
PopupScreen "Tank 1P Status" 885x425
   TrendView "Trend view_1" at 280,8 size 600x360
   TextField "Text field_4" at 20,136 size 86x22; Text 'Pressure:'
   IOField "I/O field_1" at 175,131 size 90x25; FormatPattern s999.9; Unit  mBar
      ProcessValue <- "20_TANKS_IP_DATA_RIO_01_FIRST_TANK_TANKS_PRESS"
   TextField "Text field_5" at 20,170 size 113x22; Text 'Water Level:'
   IOField "I/O field_2" at 175,165 size 90x25; FormatPattern 999.9; Unit  %
      ProcessValue <- "20_TANKS_IP_DATA_RIO_01_SECOND_TANK_BWT_LEVEL"
   TextField "Text field_6" at 20,204 size 137x22; Text 'MBG Flow Rate:'
   IOField "I/O field_3" at 175,199 size 90x25; FormatPattern 999.9; Unit  m³/hr
      ProcessValue <- "20_TANKS_IP_DATA_RIO_01_SECOND_TANK_MBG_FLOW"
   TextField "Text field_7" at 20,238 size 135x22; Text 'USD Flow Rate:'
   IOField "I/O field_4" at 175,233 size 90x25; FormatPattern 999.9; Unit  m³/hr
      ProcessValue <- "20_TANKS_IP_DATA_RIO_01_SECOND_TANK_USD_FLOW"
   TextField "Text field_8" at 20,272 size 140x22; Text 'Water pH Level:'
   IOField "I/O field_5" at 175,267 size 90x25; FormatPattern 99.9
      ProcessValue <- "20_TANKS_IP_DATA_RIO_01_SECOND_TANK_BWT_PH"
   TextField "Text field_9" at 20,306 size 143x22; Text 'Water DO Level:'
   IOField "I/O field_6" at 175,301 size 90x25; FormatPattern 99.99; Unit  mg/l
      ProcessValue <- "20_TANKS_IP_DATA_RIO_01_SECOND_TANK_BWT_DO"
   TextField "Text field_10" at 20,340 size 174x22; Text 'Water Temperature:'
   IOField "I/O field_7" at 190,335 size 75x25; FormatPattern 999.9; Unit  °C
      ProcessValue <- "20_TANKS_IP_DATA_RIO_01_SECOND_TANK_BWT_TEMP"
   Button "Button_1" at 51,5 size 219x35; TextOff 'Port Tank 1 (1P)'
      on Release: function_efd93a16("Tank 1P Status", 168, 315, -1, 0, 1)
   Button "Button_4" at 547,375 size 150x40; TextOff 'Disable Tank'; Authorization "Operate"
      on Press: function_b14e0dd5("504_Tank Grouping_DB2020_TANK ACTIV 2", 0)
   TextField "Text field_1" at 20,90 size 109x25; Text 'TIME LEFT:'
   GraphicView "Graphic view_1" at 20,46 size 245x32; Picture "Tank Manually Disabled"
   GraphicIOField "Graphic I/O field_1" at 20,46 size 245x32; PictureList "Tank Process Stage_II"
      ProcessValue <- "2110_BTCS_CNTRL_DB_BTCS_STATE"
      Visibility <- "504_Tank Grouping_DB2020_GROUP of TANK 2"
   Button "Button_2" at 4,5 size 45x35; TextOff 'Text'; PictureOff "Graphic_286"
      on Click: function_efd93a16("Tank 1P Status", 0, 0, -1, -1, 1)
   Button "Button_3" at 287,375 size 230x40; TextOff 'Text'; PictureList "Water Level Override"; Authorization "Operate"
      on Press: InvertBit("2062_Warning_Data_Water Level Override 1P")
      ProcessValue <- "2062_Warning_Data_Water Level Override 1P"
   Button "Button_5" at 27,375 size 230x40; TextOff 'Tank Shutdown Alarm'
      Visibility <- "2062_Warning_Data_Alarm Tank P1"
      ProcessValue <- "2062_Warning_Data_Water Level Override 1P"
   Button "Button_6" at 27,375 size 230x40; TextOff 'No/Low Water Level'; Authorization "Operate"
      Visibility <- "LT422 1P  TANK LEVEL ALARM_ALARM L"
      ProcessValue <- "2062_Warning_Data_Water Level Override 1P"
   IOField "I/O field_29" at 218,90 size 47x25; FormatPattern 99; Unit m
      ProcessValue <- "504_Tank Grouping_DB2020_Time Left Tank_Time Left m Tank 2"
   IOField "I/O field_8" at 173,90 size 42x25; FormatPattern 99; Unit h
      ProcessValue <- "504_Tank Grouping_DB2020_Time Left Tank_Time Left h Tank 2"
   IOField "I/O field_9" at 128,90 size 42x25; FormatPattern 99; Unit d
      ProcessValue <- "504_Tank Grouping_DB2020_Time Left Tank_Time Left d Tank 2"

PopupScreen "Tank 1S Status" 885x425
   TrendView "Trend view_1" at 280,7 size 600x360
   TextField "Text field_4" at 20,135 size 86x22; Text 'Pressure:'
   IOField "I/O field_1" at 175,130 size 90x25; FormatPattern s999.9; Unit  mBar
      ProcessValue <- "20_TANKS_IP_DATA_RIO_01_FIRST_TANK_TANKS_PRESS"
   TextField "Text field_5" at 20,169 size 113x22; Text 'Water Level:'
   IOField "I/O field_2" at 175,164 size 90x25; FormatPattern 999.9; Unit  %
      ProcessValue <- "20_TANKS_IP_DATA_RIO_01_THIRD_TANK_BWT_LEVEL"
   TextField "Text field_6" at 20,203 size 137x22; Text 'MBG Flow Rate:'
   IOField "I/O field_3" at 175,198 size 90x25; FormatPattern 999.9; Unit  m³/hr
      ProcessValue <- "20_TANKS_IP_DATA_RIO_01_THIRD_TANK_MBG_FLOW"
   TextField "Text field_7" at 20,237 size 135x22; Text 'USD Flow Rate:'
   IOField "I/O field_4" at 175,232 size 90x25; FormatPattern 999.9; Unit  m³/hr
      ProcessValue <- "20_TANKS_IP_DATA_RIO_01_THIRD_TANK_USD_FLOW"
   TextField "Text field_8" at 20,271 size 140x22; Text 'Water pH Level:'
   IOField "I/O field_5" at 175,266 size 90x25; FormatPattern 99.9
      ProcessValue <- "20_TANKS_IP_DATA_RIO_01_THIRD_TANK_BWT_PH"
   TextField "Text field_9" at 20,305 size 143x22; Text 'Water DO Level:'
   IOField "I/O field_6" at 175,300 size 90x25; FormatPattern 99.99; Unit  mg/l
      ProcessValue <- "20_TANKS_IP_DATA_RIO_01_THIRD_TANK_BWT_DO"
   TextField "Text field_10" at 20,339 size 174x22; Text 'Water Temperature:'
   IOField "I/O field_7" at 190,334 size 75x25; FormatPattern 999.9; Unit  °C
      ProcessValue <- "20_TANKS_IP_DATA_RIO_01_THIRD_TANK_BWT_TEMP"
   Button "Button_1" at 50,5 size 220x35; TextOff 'Starboard Tank 1 (1S)'
      on Release: function_efd93a16("Tank 1S Status", 168, 315, -1, 0, 1)
   Button "Button_4" at 548,375 size 150x40; TextOff 'Disable Tank'; Authorization "Operate"
      on Press: function_b14e0dd5("504_Tank Grouping_DB2020_TANK ACTIV 3", 0)
   TextField "Text field_1" at 20,90 size 109x25; Text 'TIME LEFT:'
   GraphicView "Graphic view_1" at 20,46 size 245x32; Picture "Tank Manually Disabled"
   GraphicIOField "Graphic I/O field_1" at 20,46 size 245x32; PictureList "Tank Process Stage_II"
      ProcessValue <- "2110_BTCS_CNTRL_DB_BTCS_STATE"
      Visibility <- "504_Tank Grouping_DB2020_GROUP of TANK 3"
   Button "Button_2" at 4,5 size 45x35; TextOff 'Text'; PictureOff "Graphic_286"
      on Click: function_efd93a16("Tank 1S Status", 0, 0, -1, -1, 1)
   Button "Button_3" at 287,375 size 230x40; TextOff 'Text'; PictureList "Water Level Override"; Authorization "Operate"
      on Press: InvertBit("2062_Warning_Data_Water Level Override 1S")
      ProcessValue <- "2062_Warning_Data_Water Level Override 1S"
   Button "Button_5" at 27,375 size 230x40; TextOff 'Tank Shutdown Alarm'
      Visibility <- "2062_Warning_Data_Alarm Tank S1"
   Button "Button_6" at 27,375 size 230x40; TextOff 'No/Low Water Level'; Authorization "Operate"
      Visibility <- "LT421 1S  TANK LEVEL ALARM_ALARM L"
   IOField "I/O field_29" at 218,90 size 47x25; FormatPattern 99; Unit m
      ProcessValue <- "504_Tank Grouping_DB2020_Time Left Tank_Time Left m Tank 3"
   IOField "I/O field_8" at 173,90 size 42x25; FormatPattern 99; Unit h
      ProcessValue <- "504_Tank Grouping_DB2020_Time Left Tank_Time Left h Tank 3"
   IOField "I/O field_9" at 128,90 size 42x25; FormatPattern 99; Unit d
      ProcessValue <- "504_Tank Grouping_DB2020_Time Left Tank_Time Left d Tank 3"

PopupScreen "Tank 2P Status" 885x425
   TrendView "Trend view_1" at 280,7 size 600x360
   TextField "Text field_4" at 20,135 size 86x22; Text 'Pressure:'
   IOField "I/O field_1" at 175,130 size 90x25; FormatPattern s999.9; Unit  mBar
      ProcessValue <- "20_TANKS_IP_DATA_RIO_02_FIRST_TANK_TANKS_PRESS"
   TextField "Text field_5" at 20,169 size 113x22; Text 'Water Level:'
   IOField "I/O field_2" at 175,164 size 90x25; FormatPattern 999.9; Unit  %
      ProcessValue <- "20_TANKS_IP_DATA_RIO_02_FIRST_TANK_BWT_LEVEL"
   TextField "Text field_6" at 20,203 size 137x22; Text 'MBG Flow Rate:'
   IOField "I/O field_3" at 175,198 size 90x25; FormatPattern 999.9; Unit  m³/hr
      ProcessValue <- "20_TANKS_IP_DATA_RIO_02_FIRST_TANK_MBG_FLOW"
   TextField "Text field_7" at 20,237 size 135x22; Text 'USD Flow Rate:'
   IOField "I/O field_4" at 175,232 size 90x25; FormatPattern 999.9; Unit  m³/hr
      ProcessValue <- "20_TANKS_IP_DATA_RIO_02_FIRST_TANK_USD_FLOW"
   TextField "Text field_8" at 20,271 size 140x22; Text 'Water pH Level:'
   IOField "I/O field_5" at 175,266 size 90x25; FormatPattern 99.9
      ProcessValue <- "20_TANKS_IP_DATA_RIO_02_FIRST_TANK_BWT_PH"
   TextField "Text field_9" at 20,305 size 143x22; Text 'Water DO Level:'
   IOField "I/O field_6" at 175,300 size 90x25; FormatPattern 99.99; Unit  mg/l
      ProcessValue <- "20_TANKS_IP_DATA_RIO_02_FIRST_TANK_BWT_DO"
   TextField "Text field_10" at 20,339 size 174x22; Text 'Water Temperature:'
   IOField "I/O field_7" at 190,334 size 75x25; FormatPattern 999.9; Unit  °C
      ProcessValue <- "20_TANKS_IP_DATA_RIO_02_FIRST_TANK_BWT_TEMP"
   Button "Button_4" at 545,375 size 150x40; TextOff 'Disable Tank'; Authorization "Operate"
      on Press: function_b14e0dd5("504_Tank Grouping_DB2020_TANK ACTIV 4", 0)
   Button "Button_1" at 51,5 size 219x35; TextOff 'Port Tank 2 (2P)'
      on Release: function_efd93a16("Tank 2P Status", 168, 315, -1, 0, 1)
   TextField "Text field_1" at 20,90 size 109x25; Text 'TIME LEFT:'
   GraphicView "Graphic view_1" at 20,46 size 245x32; Picture "Tank Manually Disabled"
   GraphicIOField "Graphic I/O field_1" at 20,46 size 245x32; PictureList "Tank Process Stage_II"
      ProcessValue <- "2110_BTCS_CNTRL_DB_BTCS_STATE"
      Visibility <- "504_Tank Grouping_DB2020_GROUP of TANK 4"
   Button "Button_2" at 4,5 size 45x35; TextOff 'Text'; PictureOff "Graphic_286"
      on Click: function_efd93a16("Tank 2P Status", 0, 0, -1, -1, 1)
   Button "Button_3" at 287,375 size 230x40; TextOff 'Text'; PictureList "Water Level Override"; Authorization "Operate"
      on Press: InvertBit("2062_Warning_Data_Water Level Override 2P")
      ProcessValue <- "2062_Warning_Data_Water Level Override 2P"
   Button "Button_5" at 27,375 size 230x40; TextOff 'Tank Shutdown Alarm'
      Visibility <- "2062_Warning_Data_Alarm Tank P2"
   Button "Button_6" at 27,375 size 230x40; TextOff 'No/Low Water Level'; Authorization "Operate"
      Visibility <- "FIT418_2P_ALM_ANALOG_DB_ALARM L"
   IOField "I/O field_29" at 218,90 size 47x25; FormatPattern 99; Unit m
      ProcessValue <- "504_Tank Grouping_DB2020_Time Left Tank_Time Left m Tank 4"
   IOField "I/O field_8" at 173,90 size 42x25; FormatPattern 99; Unit h
      ProcessValue <- "504_Tank Grouping_DB2020_Time Left Tank_Time Left h Tank 4"
   IOField "I/O field_9" at 128,90 size 42x25; FormatPattern 99; Unit d
      ProcessValue <- "504_Tank Grouping_DB2020_Time Left Tank_Time Left d Tank 4"

PopupScreen "Tank 2S Status" 885x425
   TrendView "Trend view_1" at 280,6 size 600x360
   TextField "Text field_4" at 20,134 size 86x22; Text 'Pressure:'
   IOField "I/O field_1" at 175,129 size 90x25; FormatPattern s999.9; Unit  mBar
      ProcessValue <- "20_TANKS_IP_DATA_RIO_02_FIRST_TANK_TANKS_PRESS"
   TextField "Text field_5" at 20,168 size 113x22; Text 'Water Level:'
   IOField "I/O field_2" at 175,163 size 90x25; FormatPattern 999.9; Unit  %
      ProcessValue <- "20_TANKS_IP_DATA_RIO_02_SECOND_TANK_BWT_LEVEL"
   TextField "Text field_6" at 20,202 size 137x22; Text 'MBG Flow Rate:'
   IOField "I/O field_3" at 175,197 size 90x25; FormatPattern 999.9; Unit  m³/hr
      ProcessValue <- "20_TANKS_IP_DATA_RIO_02_SECOND_TANK_MBG_FLOW"
   TextField "Text field_7" at 20,236 size 135x22; Text 'USD Flow Rate:'
   IOField "I/O field_4" at 175,231 size 90x25; FormatPattern 999.9; Unit  m³/hr
      ProcessValue <- "20_TANKS_IP_DATA_RIO_02_SECOND_TANK_USD_FLOW"
   TextField "Text field_8" at 20,270 size 140x22; Text 'Water pH Level:'
   IOField "I/O field_5" at 175,265 size 90x25; FormatPattern 99.9
      ProcessValue <- "20_TANKS_IP_DATA_RIO_02_SECOND_TANK_BWT_PH"
   TextField "Text field_9" at 20,304 size 143x22; Text 'Water DO Level:'
   IOField "I/O field_6" at 175,299 size 90x25; FormatPattern 99.99; Unit  mg/l
      ProcessValue <- "20_TANKS_IP_DATA_RIO_02_SECOND_TANK_BWT_DO"
   TextField "Text field_10" at 20,338 size 174x22; Text 'Water Temperature:'
   IOField "I/O field_7" at 190,333 size 75x25; FormatPattern 999.9; Unit  °C
      ProcessValue <- "20_TANKS_IP_DATA_RIO_02_SECOND_TANK_BWT_TEMP"
   Button "Button_4" at 550,375 size 150x40; TextOff 'Disable Tank'; Authorization "Operate"
      on Press: function_b14e0dd5("504_Tank Grouping_DB2020_TANK ACTIV 5", 0)
   Button "Button_1" at 50,5 size 220x35; TextOff 'Starboard Tank 2 (2S)'
      on Release: function_efd93a16("Tank 2S Status", 168, 315, -1, 0, 1)
   TextField "Text field_1" at 20,90 size 109x25; Text 'TIME LEFT:'
   GraphicView "Graphic view_1" at 20,46 size 245x32; Picture "Tank Manually Disabled"
   GraphicIOField "Graphic I/O field_1" at 20,46 size 245x32; PictureList "Tank Process Stage_II"
      ProcessValue <- "2110_BTCS_CNTRL_DB_BTCS_STATE"
      Visibility <- "504_Tank Grouping_DB2020_GROUP of TANK 5"
   Button "Button_2" at 4,5 size 45x35; TextOff 'Text'; PictureOff "Graphic_286"
      on Click: function_efd93a16("Tank 2S Status", 0, 0, -1, -1, 1)
   Button "Button_3" at 287,375 size 230x40; TextOff 'Text'; PictureList "Water Level Override"; Authorization "Operate"
      on Press: InvertBit("2062_Warning_Data_Water Level Override 2S")
      ProcessValue <- "2062_Warning_Data_Water Level Override 2S"
   Button "Button_5" at 27,375 size 230x40; TextOff 'Tank Shutdown Alarm'
      Visibility <- "2062_Warning_Data_Alarm Tank S2"
   Button "Button_6" at 27,375 size 230x40; TextOff 'No/Low Water Level'; Authorization "Operate"
      Visibility <- "LT421 2S  TANK LEVEL ALARM_ALARM L"
   IOField "I/O field_29" at 218,90 size 47x25; FormatPattern 99; Unit m
      ProcessValue <- "504_Tank Grouping_DB2020_Time Left Tank_Time Left m Tank 5"
   IOField "I/O field_8" at 173,90 size 42x25; FormatPattern 99; Unit h
      ProcessValue <- "504_Tank Grouping_DB2020_Time Left Tank_Time Left h Tank 5"
   IOField "I/O field_9" at 128,90 size 42x25; FormatPattern 99; Unit d
      ProcessValue <- "504_Tank Grouping_DB2020_Time Left Tank_Time Left d Tank 5"

PopupScreen "Tank 3P Status" 885x425
   TrendView "Trend view_1" at 280,7 size 600x360
   TextField "Text field_4" at 20,135 size 86x22; Text 'Pressure:'
   IOField "I/O field_1" at 175,130 size 90x25; FormatPattern s999.9; Unit  mBar
      ProcessValue <- "20_TANKS_IP_DATA_RIO_03_FIRST_TANK_TANKS_PRESS"
   TextField "Text field_5" at 20,169 size 113x22; Text 'Water Level:'
   IOField "I/O field_2" at 175,164 size 90x25; FormatPattern 999.9; Unit  %
      ProcessValue <- "20_TANKS_IP_DATA_RIO_03_FIRST_TANK_BWT_LEVEL"
   TextField "Text field_6" at 20,203 size 137x22; Text 'MBG Flow Rate:'
   IOField "I/O field_3" at 175,198 size 90x25; FormatPattern 999.9; Unit  m³/hr
      ProcessValue <- "20_TANKS_IP_DATA_RIO_03_FIRST_TANK_MBG_FLOW"
   TextField "Text field_7" at 20,237 size 135x22; Text 'USD Flow Rate:'
   IOField "I/O field_4" at 175,232 size 90x25; FormatPattern 999.9; Unit  m³/hr
      ProcessValue <- "20_TANKS_IP_DATA_RIO_03_FIRST_TANK_USD_FLOW"
   TextField "Text field_8" at 20,271 size 140x22; Text 'Water pH Level:'
   IOField "I/O field_5" at 175,266 size 90x25; FormatPattern 99.9
      ProcessValue <- "20_TANKS_IP_DATA_RIO_03_FIRST_TANK_BWT_PH"
   TextField "Text field_9" at 20,305 size 143x22; Text 'Water DO Level:'
   IOField "I/O field_6" at 175,300 size 90x25; FormatPattern 99.99; Unit  mg/l
      ProcessValue <- "20_TANKS_IP_DATA_RIO_03_FIRST_TANK_BWT_DO"
   TextField "Text field_10" at 20,339 size 174x22; Text 'Water Temperature:'
   IOField "I/O field_7" at 190,334 size 75x25; FormatPattern 999.9; Unit  °C
      ProcessValue <- "20_TANKS_IP_DATA_RIO_03_FIRST_TANK_BWT_TEMP"
   Button "Button_4" at 545,375 size 150x40; TextOff 'Disable Tank'; Authorization "Operate"
      on Press: function_b14e0dd5("504_Tank Grouping_DB2020_TANK ACTIV 6", 0)
   Button "Button_1" at 51,5 size 220x35; TextOff 'Port Tank 3 (3P)'
      on Release: function_efd93a16("Tank 3P Status", 168, 315, -1, 0, 1)
   TextField "Text field_1" at 20,90 size 109x25; Text 'TIME LEFT:'
   GraphicView "Graphic view_1" at 20,46 size 245x32; Picture "Tank Manually Disabled"
   GraphicIOField "Graphic I/O field_1" at 20,46 size 245x32; PictureList "Tank Process Stage_II"
      ProcessValue <- "2110_BTCS_CNTRL_DB_BTCS_STATE"
      Visibility <- "504_Tank Grouping_DB2020_GROUP of TANK 6"
   Button "Button_2" at 4,5 size 45x35; TextOff 'Text'; PictureOff "Graphic_286"
      on Click: function_efd93a16("Tank 3P Status", 0, 0, -1, -1, 1)
   Button "Button_3" at 287,375 size 230x40; TextOff 'Text'; PictureList "Water Level Override"; Authorization "Operate"
      on Press: InvertBit("2062_Warning_Data_Water Level Override 3P")
      ProcessValue <- "2062_Warning_Data_Water Level Override 3P"
   Button "Button_5" at 27,375 size 230x40; TextOff 'Tank Shutdown Alarm'
      Visibility <- "2062_Warning_Data_Alarm Tank P3"
   Button "Button_6" at 27,375 size 230x40; TextOff 'No/Low Water Level'; Authorization "Operate"
      Visibility <- "LT422 3P  TANK LEVEL ALARM_ALARM L"
   IOField "I/O field_29" at 218,90 size 47x25; FormatPattern 99; Unit m
      ProcessValue <- "504_Tank Grouping_DB2020_Time Left Tank_Time Left m Tank 6"
   IOField "I/O field_8" at 173,90 size 42x25; FormatPattern 99; Unit h
      ProcessValue <- "504_Tank Grouping_DB2020_Time Left Tank_Time Left h Tank 6"
   IOField "I/O field_9" at 128,90 size 42x25; FormatPattern 99; Unit d
      ProcessValue <- "504_Tank Grouping_DB2020_Time Left Tank_Time Left d Tank 6"

PopupScreen "Tank 3S Status" 885x425
   TrendView "Trend view_1" at 280,7 size 600x360
   TextField "Text field_4" at 20,135 size 86x22; Text 'Pressure:'
   IOField "I/O field_1" at 175,130 size 90x25; FormatPattern s999.9; Unit  mBar
      ProcessValue <- "20_TANKS_IP_DATA_RIO_03_FIRST_TANK_TANKS_PRESS"
   TextField "Text field_5" at 20,169 size 113x22; Text 'Water Level:'
   IOField "I/O field_2" at 175,164 size 90x25; FormatPattern 999.9; Unit  %
      ProcessValue <- "20_TANKS_IP_DATA_RIO_03_SECOND_TANK_BWT_LEVEL"
   TextField "Text field_6" at 20,203 size 137x22; Text 'MBG Flow Rate:'
   IOField "I/O field_3" at 175,198 size 90x25; FormatPattern 999.9; Unit  m³/hr
      ProcessValue <- "20_TANKS_IP_DATA_RIO_03_SECOND_TANK_MBG_FLOW"
   TextField "Text field_7" at 20,237 size 135x22; Text 'USD Flow Rate:'
   IOField "I/O field_4" at 175,232 size 90x25; FormatPattern 999.9; Unit  m³/hr
      ProcessValue <- "20_TANKS_IP_DATA_RIO_03_SECOND_TANK_USD_FLOW"
   TextField "Text field_8" at 20,271 size 140x22; Text 'Water pH Level:'
   IOField "I/O field_5" at 175,266 size 90x25; FormatPattern 99.9
      ProcessValue <- "20_TANKS_IP_DATA_RIO_03_SECOND_TANK_BWT_PH"
   TextField "Text field_9" at 20,305 size 143x22; Text 'Water DO Level:'
   IOField "I/O field_6" at 175,300 size 90x25; FormatPattern 99.99; Unit  mg/l
      ProcessValue <- "20_TANKS_IP_DATA_RIO_03_SECOND_TANK_BWT_DO"
   TextField "Text field_10" at 20,339 size 174x22; Text 'Water Temperature:'
   IOField "I/O field_7" at 190,334 size 75x25; FormatPattern 999.9; Unit  °C
      ProcessValue <- "20_TANKS_IP_DATA_RIO_03_SECOND_TANK_BWT_TEMP"
   Button "Button_4" at 547,375 size 150x40; TextOff 'Disable Tank'; Authorization "Operate"
      on Press: function_b14e0dd5("504_Tank Grouping_DB2020_TANK ACTIV 7", 0)
   Button "Button_1" at 51,5 size 219x35; TextOff 'Starboard Tank 3 (3S)'
      on Release: function_efd93a16("Tank 3S Status", 168, 315, -1, 0, 1)
   TextField "Text field_1" at 20,90 size 109x25; Text 'TIME LEFT:'
   GraphicView "Graphic view_1" at 20,46 size 245x32; Picture "Tank Manually Disabled"
   GraphicIOField "Graphic I/O field_1" at 20,46 size 245x32; PictureList "Tank Process Stage_II"
      ProcessValue <- "2110_BTCS_CNTRL_DB_BTCS_STATE"
      Visibility <- "504_Tank Grouping_DB2020_GROUP of TANK 7"
   Button "Button_2" at 4,5 size 45x35; TextOff 'Text'; PictureOff "Graphic_286"
      on Click: function_efd93a16("Tank 3S Status", 0, 0, -1, -1, 1)
   Button "Button_3" at 287,375 size 230x40; TextOff 'Text'; PictureList "Water Level Override"; Authorization "Operate"
      on Press: InvertBit("2062_Warning_Data_Water Level Override 3S")
      ProcessValue <- "2062_Warning_Data_Water Level Override 3S"
   Button "Button_5" at 27,375 size 230x40; TextOff 'Tank Shutdown Alarm'
      Visibility <- "2062_Warning_Data_Alarm Tank S3"
   Button "Button_6" at 27,375 size 230x40; TextOff 'No/Low Water Level'; Authorization "Operate"
      Visibility <- "LT421 3S  TANK LEVEL ALARM_ALARM L"
   IOField "I/O field_29" at 218,90 size 47x25; FormatPattern 99; Unit m
      ProcessValue <- "504_Tank Grouping_DB2020_Time Left Tank_Time Left m Tank 7"
   IOField "I/O field_8" at 173,90 size 42x25; FormatPattern 99; Unit h
      ProcessValue <- "504_Tank Grouping_DB2020_Time Left Tank_Time Left h Tank 7"
   IOField "I/O field_9" at 128,90 size 42x25; FormatPattern 99; Unit d
      ProcessValue <- "504_Tank Grouping_DB2020_Time Left Tank_Time Left d Tank 7"

PopupScreen "Tank 4P Status" 885x425
   TrendView "Trend view_1" at 280,7 size 600x360
   TextField "Text field_4" at 20,135 size 86x22; Text 'Pressure:'
   IOField "I/O field_1" at 175,130 size 90x25; FormatPattern s999.9; Unit  mBar
      ProcessValue <- "20_TANKS_IP_DATA_RIO_04_FIRST_TANK_TANKS_PRESS"
   TextField "Text field_5" at 20,169 size 113x22; Text 'Water Level:'
   IOField "I/O field_2" at 175,164 size 90x25; FormatPattern 999.9; Unit  %
      ProcessValue <- "20_TANKS_IP_DATA_RIO_04_FIRST_TANK_BWT_LEVEL"
   TextField "Text field_6" at 20,203 size 137x22; Text 'MBG Flow Rate:'
   IOField "I/O field_3" at 175,198 size 90x25; FormatPattern 999.9; Unit  m³/hr
      ProcessValue <- "20_TANKS_IP_DATA_RIO_04_FIRST_TANK_MBG_FLOW"
   TextField "Text field_7" at 20,237 size 135x22; Text 'USD Flow Rate:'
   IOField "I/O field_4" at 175,232 size 90x25; FormatPattern 999.9; Unit  m³/hr
      ProcessValue <- "20_TANKS_IP_DATA_RIO_04_FIRST_TANK_USD_FLOW"
   TextField "Text field_8" at 20,271 size 140x22; Text 'Water pH Level:'
   IOField "I/O field_5" at 175,266 size 90x25; FormatPattern 99.9
      ProcessValue <- "20_TANKS_IP_DATA_RIO_04_FIRST_TANK_BWT_PH"
   TextField "Text field_9" at 20,305 size 143x22; Text 'Water DO Level:'
   IOField "I/O field_6" at 175,300 size 90x25; FormatPattern 99.99; Unit  mg/l
      ProcessValue <- "20_TANKS_IP_DATA_RIO_04_FIRST_TANK_BWT_DO"
   TextField "Text field_10" at 20,339 size 174x22; Text 'Water Temperature:'
   IOField "I/O field_7" at 190,334 size 75x25; FormatPattern 999.9; Unit  °C
      ProcessValue <- "20_TANKS_IP_DATA_RIO_04_FIRST_TANK_BWT_TEMP"
   Button "Button_4" at 545,375 size 150x40; TextOff 'Disable Tank'; Authorization "Operate"
      on Press: function_b14e0dd5("504_Tank Grouping_DB2020_TANK ACTIV 8", 0)
   Button "Button_1" at 51,5 size 219x35; TextOff 'Port Tank 4 (4P)'
      on Release: function_efd93a16("Tank 4P Status", 168, 315, -1, 2, 1)
   TextField "Text field_1" at 20,90 size 109x25; Text 'TIME LEFT:'
   GraphicView "Graphic view_1" at 20,46 size 245x32; Picture "Tank Manually Disabled"
   GraphicIOField "Graphic I/O field_1" at 20,46 size 245x32; PictureList "Tank Process Stage_II"
      ProcessValue <- "2110_BTCS_CNTRL_DB_BTCS_STATE"
      Visibility <- "504_Tank Grouping_DB2020_GROUP of TANK 8"
   Button "Button_2" at 4,5 size 45x35; TextOff 'Text'; PictureOff "Graphic_286"
      on Click: function_efd93a16("Tank 4P Status", 0, 0, -1, -1, 1)
   Button "Button_3" at 287,375 size 230x40; TextOff 'Text'; PictureList "Water Level Override"; Authorization "Operate"
      on Press: InvertBit("2062_Warning_Data_Water Level Override 4P")
      ProcessValue <- "2062_Warning_Data_Water Level Override 4P"
   Button "Button_5" at 27,375 size 230x40; TextOff 'Tank Shutdown Alarm'
      Visibility <- "2062_Warning_Data_Alarm Tank P4"
   Button "Button_6" at 27,375 size 230x40; TextOff 'No/Low Water Level'; Authorization "Operate"
      Visibility <- "LT422 4P  TANK LEVEL ALARM_ALARM L"
   IOField "I/O field_29" at 218,90 size 47x25; FormatPattern 99; Unit m
      ProcessValue <- "504_Tank Grouping_DB2020_Time Left Tank_Time Left m Tank 8"
   IOField "I/O field_8" at 173,90 size 42x25; FormatPattern 99; Unit h
      ProcessValue <- "504_Tank Grouping_DB2020_Time Left Tank_Time Left h Tank 8"
   IOField "I/O field_9" at 128,90 size 42x25; FormatPattern 99; Unit d
      ProcessValue <- "504_Tank Grouping_DB2020_Time Left Tank_Time Left d Tank 8"

PopupScreen "Tank 4S Status" 885x425
   TrendView "Trend view_1" at 280,7 size 600x360
   TextField "Text field_4" at 20,135 size 86x22; Text 'Pressure:'
   IOField "I/O field_1" at 175,130 size 90x25; FormatPattern s999.9; Unit  mBar
      ProcessValue <- "20_TANKS_IP_DATA_RIO_04_FIRST_TANK_TANKS_PRESS"
   TextField "Text field_5" at 20,169 size 113x22; Text 'Water Level:'
   IOField "I/O field_2" at 175,164 size 90x25; FormatPattern 999.9; Unit  %
      ProcessValue <- "20_TANKS_IP_DATA_RIO_04_SECOND_TANK_BWT_LEVEL"
   TextField "Text field_6" at 20,203 size 137x22; Text 'MBG Flow Rate:'
   IOField "I/O field_3" at 175,198 size 90x25; FormatPattern 999.9; Unit  m³/hr
      ProcessValue <- "20_TANKS_IP_DATA_RIO_04_SECOND_TANK_MBG_FLOW"
   TextField "Text field_7" at 20,237 size 135x22; Text 'USD Flow Rate:'
   IOField "I/O field_4" at 175,232 size 90x25; FormatPattern 999.9; Unit  m³/hr
      ProcessValue <- "20_TANKS_IP_DATA_RIO_04_SECOND_TANK_USD_FLOW"
   TextField "Text field_8" at 20,271 size 140x22; Text 'Water pH Level:'
   IOField "I/O field_5" at 175,266 size 90x25; FormatPattern 99.9
      ProcessValue <- "20_TANKS_IP_DATA_RIO_04_SECOND_TANK_BWT_PH"
   TextField "Text field_9" at 20,305 size 143x22; Text 'Water DO Level:'
   IOField "I/O field_6" at 175,300 size 90x25; FormatPattern 99.99; Unit  mg/l
      ProcessValue <- "20_TANKS_IP_DATA_RIO_04_SECOND_TANK_BWT_DO"
   TextField "Text field_10" at 20,339 size 174x22; Text 'Water Temperature:'
   IOField "I/O field_7" at 190,334 size 75x25; FormatPattern 999.9; Unit  °C
      ProcessValue <- "20_TANKS_IP_DATA_RIO_04_SECOND_TANK_BWT_TEMP"
   Button "Button_4" at 545,375 size 150x40; TextOff 'Disable Tank'; Authorization "Operate"
      on Press: function_b14e0dd5("504_Tank Grouping_DB2020_TANK ACTIV 9", 0)
   Button "Button_1" at 50,5 size 220x35; TextOff 'Starboard Tank 4 (4S)'
      on Release: function_efd93a16("Tank 4S Status", 168, 315, -1, 2, 1)
   TextField "Text field_1" at 20,90 size 109x25; Text 'TIME LEFT:'
   GraphicView "Graphic view_1" at 20,46 size 245x32; Picture "Tank Manually Disabled"
   GraphicIOField "Graphic I/O field_1" at 20,46 size 245x32; PictureList "Tank Process Stage_II"
      ProcessValue <- "2110_BTCS_CNTRL_DB_BTCS_STATE"
      Visibility <- "504_Tank Grouping_DB2020_GROUP of TANK 9"
   Button "Button_2" at 4,5 size 45x35; TextOff 'Text'; PictureOff "Graphic_286"
      on Click: function_efd93a16("Tank 4S Status", 0, 0, -1, -1, 1)
   Button "Button_3" at 287,375 size 230x40; TextOff 'Text'; PictureList "Water Level Override"; Authorization "Operate"
      on Press: InvertBit("2062_Warning_Data_Water Level Override 4S")
      ProcessValue <- "2062_Warning_Data_Water Level Override 4S"
   Button "Button_5" at 27,375 size 230x40; TextOff 'Tank Shutdown Alarm'
      Visibility <- "2062_Warning_Data_Alarm Tank S4"
   Button "Button_6" at 27,375 size 230x40; TextOff 'No/Low Water Level'; Authorization "Operate"
      Visibility <- "LT421 4S  TANK LEVEL ALARM_ALARM L"
   IOField "I/O field_29" at 218,90 size 47x25; FormatPattern 99; Unit m
      ProcessValue <- "504_Tank Grouping_DB2020_Time Left Tank_Time Left m Tank 9"
   IOField "I/O field_8" at 173,90 size 42x25; FormatPattern 99; Unit h
      ProcessValue <- "504_Tank Grouping_DB2020_Time Left Tank_Time Left h Tank 9"
   IOField "I/O field_9" at 128,90 size 42x25; FormatPattern 99; Unit d
      ProcessValue <- "504_Tank Grouping_DB2020_Time Left Tank_Time Left d Tank 9"

PopupScreen "Tank 5P Status" 885x425
   TrendView "Trend view_1" at 280,7 size 600x360
   TextField "Text field_4" at 20,135 size 86x22; Text 'Pressure:'
   IOField "I/O field_1" at 175,130 size 90x25; FormatPattern s999.9; Unit  mBar
      ProcessValue <- "20_TANKS_IP_DATA_RIO_05_FIRST_TANK_TANKS_PRESS"
   TextField "Text field_5" at 20,169 size 113x22; Text 'Water Level:'
   IOField "I/O field_2" at 175,164 size 90x25; FormatPattern 999.9; Unit  %
      ProcessValue <- "20_TANKS_IP_DATA_RIO_05_FIRST_TANK_BWT_LEVEL"
   TextField "Text field_6" at 20,203 size 137x22; Text 'MBG Flow Rate:'
   IOField "I/O field_3" at 175,198 size 90x25; FormatPattern 999.9; Unit  m³/hr
      ProcessValue <- "20_TANKS_IP_DATA_RIO_05_FIRST_TANK_MBG_FLOW"
   TextField "Text field_7" at 20,237 size 135x22; Text 'USD Flow Rate:'
   IOField "I/O field_4" at 175,232 size 90x25; FormatPattern 999.9; Unit  m³/hr
      ProcessValue <- "20_TANKS_IP_DATA_RIO_05_FIRST_TANK_USD_FLOW"
   TextField "Text field_8" at 20,271 size 140x22; Text 'Water pH Level:'
   IOField "I/O field_5" at 175,266 size 90x25; FormatPattern 99.9
      ProcessValue <- "20_TANKS_IP_DATA_RIO_05_FIRST_TANK_BWT_PH"
   TextField "Text field_9" at 20,305 size 143x22; Text 'Water DO Level:'
   IOField "I/O field_6" at 175,300 size 90x25; FormatPattern 99.99; Unit  mg/l
      ProcessValue <- "20_TANKS_IP_DATA_RIO_05_FIRST_TANK_BWT_DO"
   TextField "Text field_10" at 20,339 size 174x22; Text 'Water Temperature:'
   IOField "I/O field_7" at 190,334 size 75x25; FormatPattern 999.9; Unit  °C
      ProcessValue <- "20_TANKS_IP_DATA_RIO_05_FIRST_TANK_BWT_TEMP"
   Button "Button_4" at 546,375 size 150x40; TextOff 'Disable Tank'; Authorization "Operate"
      on Press: function_b14e0dd5("504_Tank Grouping_DB2020_TANK ACTIV 10", 0)
   Button "Button_1" at 51,5 size 219x35; TextOff 'Port Tank 5 (5P)'
      on Release: function_efd93a16("Tank 5P Status", 168, 315, -1, 2, 1)
   TextField "Text field_1" at 20,90 size 109x25; Text 'TIME LEFT:'
   GraphicView "Graphic view_1" at 20,46 size 245x32; Picture "Tank Manually Disabled"
   GraphicIOField "Graphic I/O field_1" at 20,46 size 245x32; PictureList "Tank Process Stage_II"
      ProcessValue <- "2110_BTCS_CNTRL_DB_BTCS_STATE"
      Visibility <- "504_Tank Grouping_DB2020_GROUP of TANK 10"
   Button "Button_2" at 4,5 size 45x35; TextOff 'Text'; PictureOff "Graphic_286"
      on Click: function_efd93a16("Tank 5P Status", 0, 0, -1, -1, 1)
   Button "Button_3" at 287,375 size 230x40; TextOff 'Text'; PictureList "Water Level Override"; Authorization "Operate"
      on Press: InvertBit("2062_Warning_Data_Water Level Override 5P")
      ProcessValue <- "2062_Warning_Data_Water Level Override 5P"
   Button "Button_5" at 27,375 size 230x40; TextOff 'Tank Shutdown Alarm'
      Visibility <- "2062_Warning_Data_Alarm Tank P5"
   Button "Button_6" at 27,375 size 230x40; TextOff 'No/Low Water Level'; Authorization "Operate"
      Visibility <- "LT422 5P  TANK LEVEL ALARM_ALARM L"
   IOField "I/O field_29" at 218,90 size 47x25; FormatPattern 99; Unit m
      ProcessValue <- "504_Tank Grouping_DB2020_Time Left Tank_Time Left m Tank 10"
   IOField "I/O field_8" at 173,90 size 42x25; FormatPattern 99; Unit h
      ProcessValue <- "504_Tank Grouping_DB2020_Time Left Tank_Time Left h Tank 10"
   IOField "I/O field_9" at 128,90 size 42x25; FormatPattern 99; Unit d
      ProcessValue <- "504_Tank Grouping_DB2020_Time Left Tank_Time Left d Tank 10"

PopupScreen "Tank 5S Status" 885x425
   TrendView "Trend view_1" at 280,7 size 600x360
   TextField "Text field_4" at 20,135 size 86x22; Text 'Pressure:'
   IOField "I/O field_1" at 175,130 size 90x25; FormatPattern s999.9; Unit  mBar
      ProcessValue <- "20_TANKS_IP_DATA_RIO_05_FIRST_TANK_TANKS_PRESS"
   TextField "Text field_5" at 20,169 size 113x22; Text 'Water Level:'
   IOField "I/O field_2" at 175,164 size 90x25; FormatPattern 999.9; Unit  %
      ProcessValue <- "20_TANKS_IP_DATA_RIO_05_SECOND_TANK_BWT_LEVEL"
   TextField "Text field_6" at 20,203 size 137x22; Text 'MBG Flow Rate:'
   IOField "I/O field_3" at 175,198 size 90x25; FormatPattern 999.9; Unit  m³/hr
      ProcessValue <- "20_TANKS_IP_DATA_RIO_05_SECOND_TANK_MBG_FLOW"
   TextField "Text field_7" at 20,237 size 135x22; Text 'USD Flow Rate:'
   IOField "I/O field_4" at 175,232 size 90x25; FormatPattern 999.9; Unit  m³/hr
      ProcessValue <- "20_TANKS_IP_DATA_RIO_05_SECOND_TANK_USD_FLOW"
   TextField "Text field_8" at 20,271 size 140x22; Text 'Water pH Level:'
   IOField "I/O field_5" at 175,266 size 90x25; FormatPattern 99.9
      ProcessValue <- "20_TANKS_IP_DATA_RIO_05_SECOND_TANK_BWT_PH"
   TextField "Text field_9" at 20,305 size 143x22; Text 'Water DO Level:'
   IOField "I/O field_6" at 175,300 size 90x25; FormatPattern 99.99; Unit  mg/l
      ProcessValue <- "20_TANKS_IP_DATA_RIO_05_SECOND_TANK_BWT_DO"
   TextField "Text field_10" at 20,339 size 174x22; Text 'Water Temperature:'
   IOField "I/O field_7" at 190,334 size 75x25; FormatPattern 999.9; Unit  °C
      ProcessValue <- "20_TANKS_IP_DATA_RIO_05_SECOND_TANK_BWT_TEMP"
   Button "Button_4" at 550,375 size 150x40; TextOff 'Disable Tank'; Authorization "Operate"
      on Press: function_b14e0dd5("504_Tank Grouping_DB2020_TANK ACTIV 11", 0)
   Button "Button_1" at 50,5 size 220x35; TextOff 'Starboard Tank 5 (5S)'
      on Release: function_efd93a16("Tank 5S Status", 168, 315, -1, 2, 1)
   TextField "Text field_1" at 20,90 size 109x25; Text 'TIME LEFT:'
   GraphicView "Graphic view_1" at 20,46 size 245x32; Picture "Tank Manually Disabled"
   GraphicIOField "Graphic I/O field_1" at 20,46 size 245x32; PictureList "Tank Process Stage_II"
      ProcessValue <- "2110_BTCS_CNTRL_DB_BTCS_STATE"
      Visibility <- "504_Tank Grouping_DB2020_GROUP of TANK 11"
   Button "Button_2" at 4,5 size 45x35; TextOff 'Text'; PictureOff "Graphic_286"
      on Click: function_efd93a16("Tank 5S Status", 0, 0, -1, -1, 1)
   Button "Button_3" at 287,375 size 230x40; TextOff 'Text'; PictureList "Water Level Override"; Authorization "Operate"
      on Press: InvertBit("2062_Warning_Data_Water Level Override 5S")
      ProcessValue <- "2062_Warning_Data_Water Level Override 5S"
   Button "Button_5" at 27,375 size 230x40; TextOff 'Tank Shutdown Alarm'
      Visibility <- "2062_Warning_Data_Alarm Tank S5"
   Button "Button_6" at 27,375 size 230x40; TextOff 'No/Low Water Level'; Authorization "Operate"
      Visibility <- "LT421 5S  TANK LEVEL ALARM_ALARM L"
   IOField "I/O field_29" at 218,90 size 47x25; FormatPattern 99; Unit m
      ProcessValue <- "504_Tank Grouping_DB2020_Time Left Tank_Time Left m Tank 11"
   IOField "I/O field_8" at 173,90 size 42x25; FormatPattern 99; Unit h
      ProcessValue <- "504_Tank Grouping_DB2020_Time Left Tank_Time Left h Tank 11"
   IOField "I/O field_9" at 128,90 size 42x25; FormatPattern 99; Unit d
      ProcessValue <- "504_Tank Grouping_DB2020_Time Left Tank_Time Left d Tank 11"

PopupScreen "Tank 6P Status" 885x425
   TrendView "Trend view_1" at 280,7 size 600x360
   TextField "Text field_4" at 20,135 size 86x22; Text 'Pressure:'
   IOField "I/O field_1" at 175,130 size 90x25; FormatPattern s999.9; Unit  mBar
      ProcessValue <- "20_TANKS_IP_DATA_RIO_06_FIRST_TANK_TANKS_PRESS"
   TextField "Text field_5" at 20,169 size 113x22; Text 'Water Level:'
   IOField "I/O field_2" at 175,164 size 90x25; FormatPattern 999.9; Unit  %
      ProcessValue <- "20_TANKS_IP_DATA_RIO_06_FIRST_TANK_BWT_LEVEL"
   TextField "Text field_6" at 20,203 size 137x22; Text 'MBG Flow Rate:'
   IOField "I/O field_3" at 175,198 size 90x25; FormatPattern 999.9; Unit  m³/hr
      ProcessValue <- "20_TANKS_IP_DATA_RIO_06_FIRST_TANK_MBG_FLOW"
   TextField "Text field_7" at 20,237 size 135x22; Text 'USD Flow Rate:'
   IOField "I/O field_4" at 175,232 size 90x25; FormatPattern 999.9; Unit  m³/hr
      ProcessValue <- "20_TANKS_IP_DATA_RIO_06_FIRST_TANK_USD_FLOW"
   TextField "Text field_8" at 20,271 size 140x22; Text 'Water pH Level:'
   IOField "I/O field_5" at 175,266 size 90x25; FormatPattern 99.9
      ProcessValue <- "20_TANKS_IP_DATA_RIO_06_FIRST_TANK_BWT_PH"
   TextField "Text field_9" at 20,305 size 143x22; Text 'Water DO Level:'
   IOField "I/O field_6" at 175,300 size 90x25; FormatPattern 99.99; Unit  mg/l
      ProcessValue <- "20_TANKS_IP_DATA_RIO_06_FIRST_TANK_BWT_DO"
   TextField "Text field_10" at 20,339 size 174x22; Text 'Water Temperature:'
   IOField "I/O field_7" at 190,334 size 75x25; FormatPattern 999.9; Unit  °C
      ProcessValue <- "20_TANKS_IP_DATA_RIO_06_FIRST_TANK_BWT_TEMP"
   Button "Button_4" at 542,374 size 150x40; TextOff 'Disable Tank'; Authorization "Operate"
      on Press: function_b14e0dd5("504_Tank Grouping_DB2020_TANK ACTIV 12", 0)
   Button "Button_1" at 51,5 size 219x35; TextOff 'Port Tank 6 (6P)'
      on Release: function_efd93a16("Tank 6P Status", 168, 315, -1, 2, 1)
   TextField "Text field_1" at 20,90 size 109x25; Text 'TIME LEFT:'
   GraphicView "Graphic view_1" at 20,46 size 245x32; Picture "Tank Manually Disabled"
   GraphicIOField "Graphic I/O field_1" at 20,46 size 245x32; PictureList "Tank Process Stage_II"
      ProcessValue <- "2110_BTCS_CNTRL_DB_BTCS_STATE"
      Visibility <- "504_Tank Grouping_DB2020_GROUP of TANK 12"
   Button "Button_2" at 4,5 size 45x35; TextOff 'Text'; PictureOff "Graphic_286"
      on Click: function_efd93a16("Tank 6P Status", 0, 0, -1, -1, 1)
   Button "Button_3" at 287,375 size 230x40; TextOff 'Text'; PictureList "Water Level Override"; Authorization "Operate"
      on Press: InvertBit("2062_Warning_Data_Water Level Override 6P")
      ProcessValue <- "2062_Warning_Data_Water Level Override 6P"
   Button "Button_5" at 27,375 size 230x40; TextOff 'Tank Shutdown Alarm'
      Visibility <- "2062_Warning_Data_Alarm Tank P6"
   Button "Button_6" at 27,375 size 230x40; TextOff 'No/Low Water Level'; Authorization "Operate"
      Visibility <- "LT422 6P  TANK LEVEL ALARM_ALARM L"
   IOField "I/O field_29" at 218,90 size 47x25; FormatPattern 99; Unit m
      ProcessValue <- "504_Tank Grouping_DB2020_Time Left Tank_Time Left m Tank 12"
   IOField "I/O field_8" at 173,90 size 42x25; FormatPattern 99; Unit h
      ProcessValue <- "504_Tank Grouping_DB2020_Time Left Tank_Time Left h Tank 12"
   IOField "I/O field_9" at 128,90 size 42x25; FormatPattern 99; Unit d
      ProcessValue <- "504_Tank Grouping_DB2020_Time Left Tank_Time Left d Tank 12"

PopupScreen "Tank 6S Status" 885x425
   TrendView "Trend view_1" at 280,7 size 600x360
   TextField "Text field_4" at 20,135 size 86x22; Text 'Pressure:'
   IOField "I/O field_1" at 175,130 size 90x25; FormatPattern s999.9; Unit  mBar
      ProcessValue <- "20_TANKS_IP_DATA_RIO_06_FIRST_TANK_TANKS_PRESS"
   TextField "Text field_5" at 20,169 size 113x22; Text 'Water Level:'
   IOField "I/O field_2" at 175,164 size 90x25; FormatPattern 999.9; Unit  %
      ProcessValue <- "20_TANKS_IP_DATA_RIO_06_SECOND_TANK_BWT_LEVEL"
   TextField "Text field_6" at 20,203 size 137x22; Text 'MBG Flow Rate:'
   IOField "I/O field_3" at 175,198 size 90x25; FormatPattern 999.9; Unit  m³/hr
      ProcessValue <- "20_TANKS_IP_DATA_RIO_06_SECOND_TANK_MBG_FLOW"
   TextField "Text field_7" at 20,237 size 135x22; Text 'USD Flow Rate:'
   IOField "I/O field_4" at 175,232 size 90x25; FormatPattern 999.9; Unit  m³/hr
      ProcessValue <- "20_TANKS_IP_DATA_RIO_06_SECOND_TANK_USD_FLOW"
   TextField "Text field_8" at 20,271 size 140x22; Text 'Water pH Level:'
   IOField "I/O field_5" at 175,266 size 90x25; FormatPattern 99.9
      ProcessValue <- "20_TANKS_IP_DATA_RIO_06_SECOND_TANK_BWT_PH"
   TextField "Text field_9" at 20,305 size 143x22; Text 'Water DO Level:'
   IOField "I/O field_6" at 175,300 size 90x25; FormatPattern 99.99; Unit  mg/l
      ProcessValue <- "20_TANKS_IP_DATA_RIO_06_SECOND_TANK_BWT_DO"
   TextField "Text field_10" at 20,339 size 174x22; Text 'Water Temperature:'
   IOField "I/O field_7" at 190,334 size 75x25; FormatPattern 999.9; Unit  °C
      ProcessValue <- "20_TANKS_IP_DATA_RIO_06_SECOND_TANK_BWT_TEMP"
   Button "Button_4" at 545,377 size 150x40; TextOff 'Disable Tank'; Authorization "Operate"
      on Press: function_b14e0dd5("504_Tank Grouping_DB2020_TANK ACTIV 13", 0)
   Button "Button_1" at 51,5 size 219x35; TextOff 'Starboard Tank 6 (6S)'
      on Release: function_efd93a16("Tank 6S Status", 168, 315, -1, 2, 1)
   TextField "Text field_1" at 20,90 size 109x25; Text 'TIME LEFT:'
   GraphicView "Graphic view_1" at 20,46 size 245x32; Picture "Tank Manually Disabled"
   GraphicIOField "Graphic I/O field_1" at 20,46 size 245x32; PictureList "Tank Process Stage_II"
      ProcessValue <- "2110_BTCS_CNTRL_DB_BTCS_STATE"
      Visibility <- "504_Tank Grouping_DB2020_GROUP of TANK 13"
   Button "Button_2" at 4,5 size 45x35; TextOff 'Text'; PictureOff "Graphic_286"
      on Click: function_efd93a16("Tank 6S Status", 0, 0, -1, -1, 1)
   Button "Button_3" at 287,375 size 230x40; TextOff 'Text'; PictureList "Water Level Override"; Authorization "Operate"
      on Press: InvertBit("2062_Warning_Data_Water Level Override 6S")
      ProcessValue <- "2062_Warning_Data_Water Level Override 6S"
   Button "Button_5" at 27,375 size 230x40; TextOff 'Tank Shutdown Alarm'
      Visibility <- "2062_Warning_Data_Alarm Tank S6"
   Button "Button_6" at 27,375 size 230x40; TextOff 'No/Low Water Level'; Authorization "Operate"
      Visibility <- "LT421 6S  TANK LEVEL ALARM_ALARM L"
   IOField "I/O field_29" at 218,90 size 47x25; FormatPattern 99; Unit m
      ProcessValue <- "504_Tank Grouping_DB2020_Time Left Tank_Time Left m Tank 13"
   IOField "I/O field_8" at 173,90 size 42x25; FormatPattern 99; Unit h
      ProcessValue <- "504_Tank Grouping_DB2020_Time Left Tank_Time Left h Tank 13"
   IOField "I/O field_9" at 128,90 size 42x25; FormatPattern 99; Unit d
      ProcessValue <- "504_Tank Grouping_DB2020_Time Left Tank_Time Left d Tank 13"

PopupScreen "Tank AP Status" 885x425
   TrendView "Trend view_1" at 280,7 size 600x360
   TextField "Text field_4" at 20,135 size 86x22; Text 'Pressure:'
   IOField "I/O field_1" at 175,130 size 90x25; FormatPattern s999.9; Unit  mBar
      ProcessValue <- "20_TANKS_IP_DATA_RIO_07_FIRST_TANK_TANKS_PRESS"
   TextField "Text field_5" at 20,169 size 113x22; Text 'Water Level:'
   IOField "I/O field_2" at 175,164 size 90x25; FormatPattern 999.9; Unit  %
      ProcessValue <- "20_TANKS_IP_DATA_RIO_07_FIRST_TANK_BWT_LEVEL"
   TextField "Text field_6" at 20,203 size 137x22; Text 'MBG Flow Rate:'
   IOField "I/O field_3" at 175,198 size 90x25; FormatPattern 999.9; Unit  m³/hr
      ProcessValue <- "20_TANKS_IP_DATA_RIO_07_FIRST_TANK_MBG_FLOW"
   TextField "Text field_7" at 20,237 size 135x22; Text 'USD Flow Rate:'
   IOField "I/O field_4" at 175,232 size 90x25; FormatPattern 999.9; Unit  m³/hr
      ProcessValue <- "20_TANKS_IP_DATA_RIO_07_FIRST_TANK_USD_FLOW"
   TextField "Text field_8" at 20,271 size 140x22; Text 'Water pH Level:'
   IOField "I/O field_5" at 175,266 size 90x25; FormatPattern 99.9
      ProcessValue <- "20_TANKS_IP_DATA_RIO_07_FIRST_TANK_BWT_PH"
   TextField "Text field_9" at 20,305 size 143x22; Text 'Water DO Level:'
   IOField "I/O field_6" at 175,300 size 90x25; FormatPattern 99.99; Unit  mg/l
      ProcessValue <- "20_TANKS_IP_DATA_RIO_07_FIRST_TANK_BWT_DO"
   TextField "Text field_10" at 20,339 size 174x22; Text 'Water Temperature:'
   IOField "I/O field_7" at 190,334 size 75x25; FormatPattern 999.9; Unit  °C
      ProcessValue <- "20_TANKS_IP_DATA_RIO_07_FIRST_TANK_BWT_TEMP"
   Button "Button_4" at 538,375 size 150x40; TextOff 'Disable Tank'; Authorization "Operate"
      on Press: function_b14e0dd5("504_Tank Grouping_DB2020_TANK ACTIV 14", 0)
   Button "Button_1" at 51,5 size 219x35; TextOff 'Aft Peak Tank (APT)'
      on Release: function_efd93a16("Tank AP Status", 168, 315, -1, 2, 1)
   TextField "Text field_1" at 20,90 size 109x25; Text 'TIME LEFT:'
   GraphicView "Graphic view_1" at 20,46 size 245x32; Picture "Tank Manually Disabled"
   GraphicIOField "Graphic I/O field_1" at 20,46 size 245x32; PictureList "Tank Process Stage_II"
      ProcessValue <- "2110_BTCS_CNTRL_DB_BTCS_STATE"
      Visibility <- "504_Tank Grouping_DB2020_GROUP of TANK 14"
   Button "Button_2" at 4,5 size 45x35; TextOff 'Text'; PictureOff "Graphic_286"
      on Click: function_efd93a16("Tank AP Status", 0, 0, -1, -1, 1)
   Button "Button_3" at 287,375 size 230x40; TextOff 'Text'; PictureList "Water Level Override"; Authorization "Operate"
      on Press: InvertBit("2062_Warning_Data_Water Level Override APT")
      ProcessValue <- "2062_Warning_Data_Water Level Override APT"
   Button "Button_5" at 27,375 size 230x40; TextOff 'Tank Shutdown Alarm'
      Visibility <- "2062_Warning_Data_Alarm Tank APT"
   Button "Button_6" at 27,375 size 230x40; TextOff 'No/Low Water Level'; Authorization "Operate"
      Visibility <- "LT422 APT  TANK LEVEL ALARM_ALARM L"
   IOField "I/O field_29" at 218,90 size 47x25; FormatPattern 99; Unit m
      ProcessValue <- "504_Tank Grouping_DB2020_Time Left Tank_Time Left m Tank 14"
   IOField "I/O field_8" at 173,90 size 42x25; FormatPattern 99; Unit h
      ProcessValue <- "504_Tank Grouping_DB2020_Time Left Tank_Time Left h Tank 14"
   IOField "I/O field_9" at 128,90 size 42x25; FormatPattern 99; Unit d
      ProcessValue <- "504_Tank Grouping_DB2020_Time Left Tank_Time Left d Tank 14"

PopupScreen "Tank FP Status" 885x425
   TrendView "Trend view_1" at 280,7 size 600x360
   TextField "Text field_1" at 20,90 size 109x25; Text 'TIME LEFT:'
   TextField "Text field_4" at 20,135 size 86x22; Text 'Pressure:'
   IOField "I/O field_1" at 175,130 size 90x25; FormatPattern s999.9; Unit  mBar
      ProcessValue <- "20_TANKS_IP_DATA_RIO_01_FIRST_TANK_TANKS_PRESS"
   TextField "Text field_5" at 20,169 size 113x22; Text 'Water Level:'
   IOField "I/O field_2" at 175,164 size 90x25; FormatPattern 999.9; Unit  %
      ProcessValue <- "20_TANKS_IP_DATA_RIO_01_FIRST_TANK_BWT_LEVEL"
   TextField "Text field_6" at 20,203 size 137x22; Text 'MBG Flow Rate:'
   IOField "I/O field_3" at 175,198 size 90x25; FormatPattern 999.9; Unit  m³/hr
      ProcessValue <- "20_TANKS_IP_DATA_RIO_01_FIRST_TANK_MBG_FLOW"
   TextField "Text field_7" at 20,237 size 135x22; Text 'USD Flow Rate:'
   IOField "I/O field_4" at 175,232 size 90x25; FormatPattern 999.9; Unit  m³/hr
      ProcessValue <- "20_TANKS_IP_DATA_RIO_01_FIRST_TANK_USD_FLOW"
   TextField "Text field_8" at 20,271 size 140x22; Text 'Water pH Level:'
   IOField "I/O field_5" at 175,266 size 90x25; FormatPattern 99.9
      ProcessValue <- "20_TANKS_IP_DATA_RIO_01_FIRST_TANK_BWT_PH"
   TextField "Text field_9" at 20,305 size 143x22; Text 'Water DO Level:'
   IOField "I/O field_6" at 175,300 size 90x25; FormatPattern 99.99; Unit  mg/l
      ProcessValue <- "20_TANKS_IP_DATA_RIO_01_FIRST_TANK_BWT_DO"
   TextField "Text field_10" at 20,339 size 174x22; Text 'Water Temperature:'
   IOField "I/O field_7" at 190,334 size 75x25; FormatPattern 999.9; Unit  °C
      ProcessValue <- "20_TANKS_IP_DATA_RIO_01_FIRST_TANK_BWT_TEMP"
   IOField "I/O field_29" at 218,90 size 47x25; FormatPattern 99; Unit m
      ProcessValue <- "504_Tank Grouping_DB2020_Time Left Tank_Time Left m Tank 1"
   Button "Button_2" at 712,375 size 150x40; TextOff 'Reset Tank'
      Visibility <- "AlwaysTRUE"
   Button "Button_3" at 287,375 size 230x40; TextOff 'Text'; PictureList "Water Level Override"; Authorization "Operate"
      on Press: InvertBit("2062_Warning_Data_Water Level Override FPT")
      ProcessValue <- "2062_Warning_Data_Water Level Override FPT"
   Button "Button_4" at 539,375 size 150x40; TextOff 'Disable Tank'; Authorization "Operate"
      on Press: function_b14e0dd5("504_Tank Grouping_DB2020_TANK ACTIV 1", 0)
   Button "Button_5" at 27,375 size 230x40; TextOff 'Tank Shutdown Alarm'
      Visibility <- "2062_Warning_Data_Alarm Tank FPT"
      ProcessValue <- "2062_Warning_Data_Water Level Override FPT"
   Button "Button_6" at 27,375 size 230x40; TextOff 'No/Low Water Level'
      Visibility <- "LT422 FPT  TANK LEVEL ALARM_ALARM L"
      ProcessValue <- "2062_Warning_Data_Water Level Override FPT"
   GraphicView "Graphic view_1" at 20,46 size 245x32; Picture "Tank Manually Disabled"
   Button "Button_1" at 51,5 size 219x35; TextOff 'Fore Peak Tank (FPT)'
   GraphicIOField "Graphic I/O field_1" at 20,46 size 245x32; PictureList "Tank Process Stage_II"
      ProcessValue <- "2110_BTCS_CNTRL_DB_BTCS_STATE"
      Visibility <- "504_Tank Grouping_DB2020_GROUP of TANK 1"
   Button "Button_7" at 4,5 size 45x35; TextOff 'Text'; PictureOff "Graphic_286"
      on Click: function_efd93a16("Tank FP Status", 0, 0, -1, -1, 1)
   IOField "I/O field_8" at 173,90 size 42x25; FormatPattern 99; Unit h
      ProcessValue <- "504_Tank Grouping_DB2020_Time Left Tank_Time Left h Tank 1"
   IOField "I/O field_9" at 128,90 size 42x25; FormatPattern 99; Unit d
      ProcessValue <- "504_Tank Grouping_DB2020_Time Left Tank_Time Left d Tank 1"

